(* Logix 5000 project; controller MV vendor 1 type 14 code 217 rev 31.11; software revision 31.00; part 41 of 53 *)
(* tags used below, declared in another part *)
   CurrentTime : DateTime;
   MV_B100 : INT[255];   // AT FLAGS
   MV_DayOfWeek : DINT;
   MV_F8 : REAL[20];
   MV_GasAvailable : BOOL;
   MV_MV10_CV1 : PlantItem;   // MV10_CV1
   MV_MV11_CV1 : PlantItem;   // MV11_CV1
   MV_MV12_CV1 : PlantItem;   // MV12_CV1
   MV_MV13_CV1 : PlantItem;   // MV13_CV1
   MV_MV14_CV1 : PlantItem;   // MV14_CV1
   MV_MV15_CV1 : PlantItem;   // MV15_CV1
   MV_MV16_CV1 : PlantItem;   // MV16_CV1
   MV_MV17_CV1 : PlantItem;   // MV17_CV1
   MV_MV18_CV1 : PlantItem;   // MV18_CV1
   MV_MV19_CV1 : PlantItem;   // MV19_CV1
   MV_MV1_CV1 : PlantItem;   // MV1_CV1
   MV_MV20_CV1 : PlantItem;   // MV20_CV1
   MV_MV21_CV1 : PlantItem;   // MV21_CV1
   MV_MV22_CV1 : PlantItem;   // MV22_CV1
   MV_MV23_CV1 : PlantItem;   // MV23_CV1
   MV_MV2_CV1 : PlantItem;   // MV2_CV1
   MV_MV30_CV1 : PlantItem;   // MV30_CV1
   MV_MV31_CV1 : PlantItem;   // MV31_CV1
   MV_MV32_CV1 : PlantItem;   // MV32_CV1
   MV_MV33_CV1 : PlantItem;   // MV33_CV1
   MV_MV34_CV1 : PlantItem;   // MV34_CV1
   MV_MV35_CV1 : PlantItem;   // MV35_CV1
   MV_MV36_AV01 : PlantItem;   // MV36_AV01
   MV_MV37_AV01 : PlantItem;   // MV37_AV01
   MV_MV38_AV01 : PlantItem;   // MV38_AV01
   MV_MV39_AV01 : PlantItem;   // MV39_AV01
   MV_MV3_CV1 : PlantItem;   // MV3_CV1
   MV_MV40_AV01 : PlantItem;   // MV40_AV01
   MV_MV41_AV01 : PlantItem;   // MV41_AV01
   MV_MV42_AV01 : PlantItem;   // MV42_AV01
   MV_MV43_AV01 : PlantItem;   // MV43_AV01
   MV_MV44_AV01 : PlantItem;   // MV44_AV01
   MV_MV45_AV01 : PlantItem;   // MV45_AV01
   MV_MV46_AV01 : PlantItem;   // MV46_AV01
   MV_MV47_AV01 : PlantItem;   // MV47_AV01
   MV_MV4_CV1 : PlantItem;   // MV4_CV1
   MV_MV5_CV1 : PlantItem;   // MV5_CV1
   MV_MV6_CV1 : PlantItem;   // MV6_CV1
   MV_MV7_CV1 : PlantItem;   // MV7_CV1
   MV_MV8_CV1 : PlantItem;   // MV8_CV1
   MV_MV9_CV1 : PlantItem;   // MV9_CV1
   MV_N101 : INT[255];   // AT INT Fermentation control integer workspace
   MV_N110 : INT[255];   // MV DATA 0 CURRENT FV DATA
   MV_N111 : INT[50];   // MV 1, CURRENT FV DATA
   MV_N112 : INT[50];   // MV 2, CURRENT FV DATA
   MV_N113 : INT[50];   // MV 3, CURRENT FV DATA
   MV_N114 : INT[50];   // MV 4, CURRENT FV DATA
   MV_N115 : INT[50];   // MV 5, CURRENT FV DATA
   MV_N116 : INT[50];   // MV 6, CURRENT FV DATA
   MV_N117 : INT[50];   // MV 7, CURRENT FV DATA
   MV_N118 : INT[50];   // MV 8, CURRENT FV DATA
   MV_N119 : INT[50];   // MV 9, CURRENT FV DATA
   MV_N12 : INT[255];   // SYS_PARMS System Parameter Fil e
   MV_N120 : INT[50];   // MV 10, CURRENT FV DATA
   MV_N121 : INT[50];   // MV 11, CURRENT FV DATA
   MV_N122 : INT[50];   // MV 12, CURRENT FV DATA
   MV_N123 : INT[50];   // MV 13, CURRENT FV DATA
   MV_N124 : INT[50];   // MV 14, CURRENT FV DATA
   MV_N125 : INT[50];   // MV 15, CURRENT FV DATA
   MV_N126 : INT[50];   // MV 16, CURRENT FV DATA
   MV_N127 : INT[50];   // MV 17, CURRENT FV DATA
   MV_N128 : INT[50];   // MV 18, CURRENT FV DATA
   MV_N129 : INT[50];   // MV 19, CURRENT FV DATA
   MV_N130 : INT[50];   // MV 30, CURRENT FV DATA
   MV_N131 : INT[50];   // MV 31, CURRENT FV DATA
   MV_N132 : INT[50];   // MV 32, CURRENT FV DATA
   MV_N133 : INT[50];   // MV 33, CURRENT FV DATA
   MV_N134 : INT[50];   // MV 34, CURRENT FV DATA
   MV_N135 : INT[50];   // MV 35, CURRENT FV DATA
   MV_N136 : INT[50];   // MV 20, CURRENT FV DATA
   MV_N137 : INT[50];   // MV 21, CURRENT FV DATA
   MV_N138 : INT[50];   // MV 22, CURRENT FV DATA
   MV_N139 : INT[50];   // MV 23, CURRENT FV DATA
   MV_N140 : INT[50];   // MV 36, CURRENT FV DATA
   MV_N141 : INT[50];   // MV 37, CURRENT FV DATA
   MV_N142 : INT[50];   // MV 38, CURRENT FV DATA
   MV_N143 : INT[50];   // MV 39, CURRENT FV DATA
   MV_N144 : INT[50];   // MV 40, CURRENT FV DATA
   MV_N145 : INT[50];   // MV 41, CURRENT FV DATA
   MV_N146 : INT[50];   // MV 42, CURRENT FV DATA
   MV_N147 : INT[50];   // MV 43, CURRENT FV DATA
   MV_N148 : INT[50];   // MV 44, CURRENT FV DATA
   MV_N149 : INT[50];   // MV 45, CURRENT FV DATA
   MV_N150 : INT[50];   // MV 36, CURRENT FV DATA
   MV_N151 : INT[50];   // MV 47, CURRENT FV DATA
   MV_SFile : INT[255];   // SLC Equivalent System File, So Original Code Can Remain
   temp : INT;
(* MV_Common, continued *)

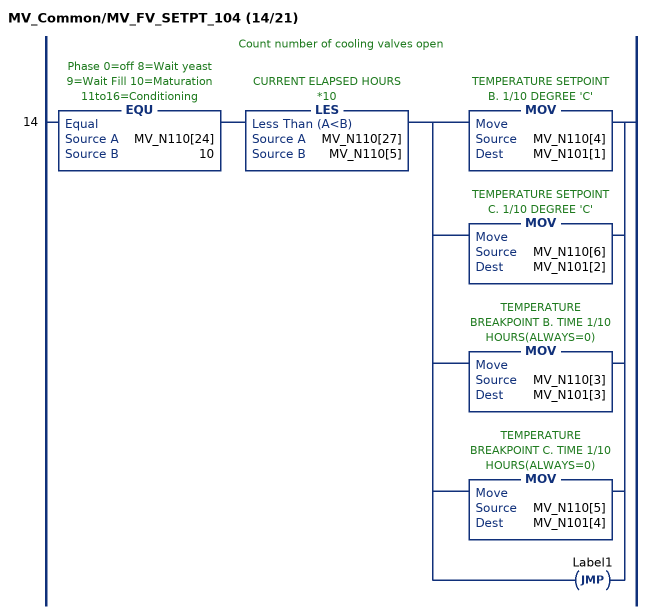
   [picture p954: MV_Common/MV_FV_SETPT_104 rungs 14-14]
   // Count number of cooling valves open
   14: EQU(MV_N110[24],10)LES(MV_N110[27],MV_N110[5])[MOV(MV_N110[4],MV_N101[1]) ,MOV(MV_N110[6],MV_N101[2]) ,MOV(MV_N110[3],MV_N101[3]) ,MOV(MV_N110[5],MV_N101[4]) ,JMP(Label1) ];
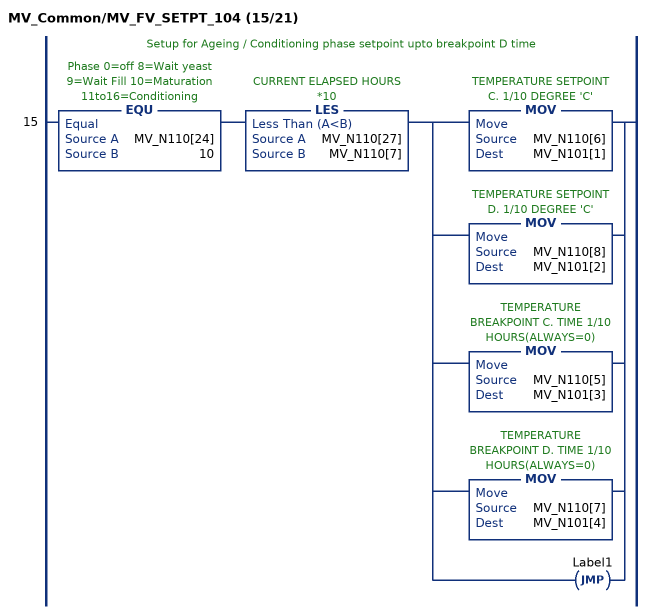
   // Setup for Ageing / Conditioning phase setpoint upto breakpoint D time
   15: EQU(MV_N110[24],10)LES(MV_N110[27],MV_N110[7])[MOV(MV_N110[6],MV_N101[1]) ,MOV(MV_N110[8],MV_N101[2]) ,MOV(MV_N110[5],MV_N101[3]) ,MOV(MV_N110[7],MV_N101[4]) ,JMP(Label1) ];
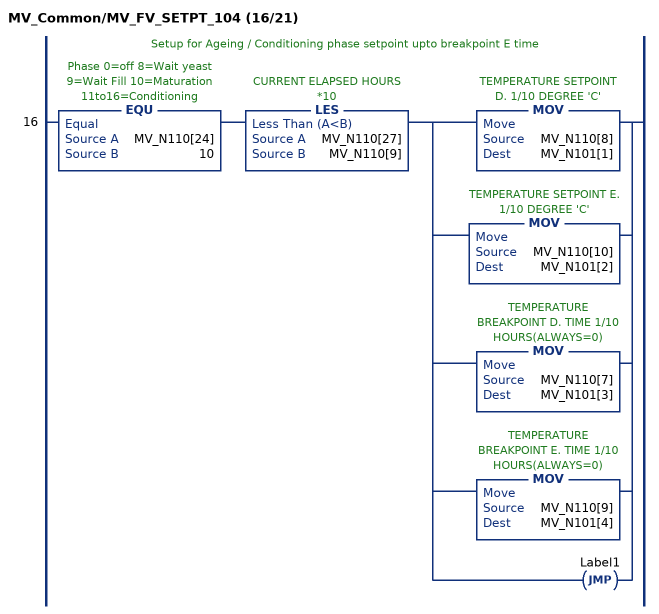
   // Setup for Ageing / Conditioning phase setpoint upto breakpoint E time
   16: EQU(MV_N110[24],10)LES(MV_N110[27],MV_N110[9])[MOV(MV_N110[8],MV_N101[1]) ,MOV(MV_N110[10],MV_N101[2]) ,MOV(MV_N110[7],MV_N101[3]) ,MOV(MV_N110[9],MV_N101[4]) ,JMP(Label1) ];
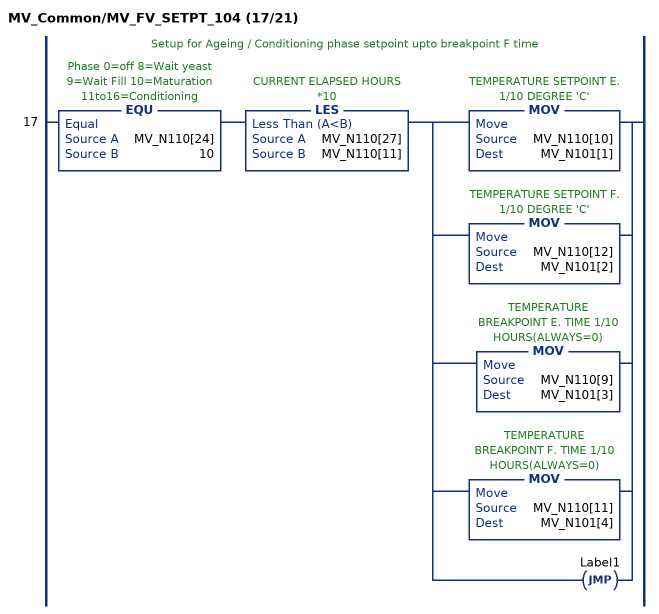
   // Setup for Ageing / Conditioning phase setpoint upto breakpoint F time
   17: EQU(MV_N110[24],10)LES(MV_N110[27],MV_N110[11])[MOV(MV_N110[10],MV_N101[1]) ,MOV(MV_N110[12],MV_N101[2]) ,MOV(MV_N110[9],MV_N101[3]) ,MOV(MV_N110[11],MV_N101[4]) ,JMP(Label1) ];
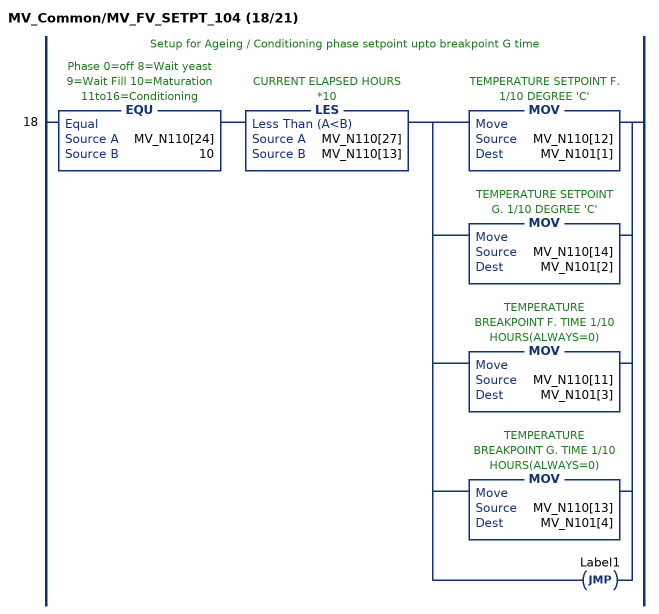
   // Setup for Ageing / Conditioning phase setpoint upto breakpoint G time
   18: EQU(MV_N110[24],10)LES(MV_N110[27],MV_N110[13])[MOV(MV_N110[12],MV_N101[1]) ,MOV(MV_N110[14],MV_N101[2]) ,MOV(MV_N110[11],MV_N101[3]) ,MOV(MV_N110[13],MV_N101[4]) ,JMP(Label1) ];
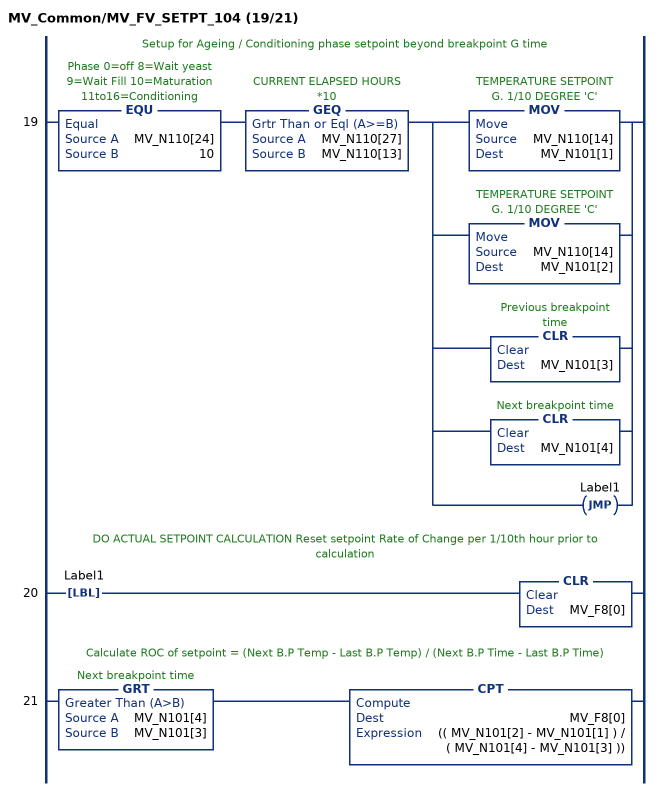
   // Setup for Ageing / Conditioning phase setpoint beyond breakpoint G time
   19: EQU(MV_N110[24],10)GEQ(MV_N110[27],MV_N110[13])[MOV(MV_N110[14],MV_N101[1]) ,MOV(MV_N110[14],MV_N101[2]) ,CLR(MV_N101[3]) ,CLR(MV_N101[4]) ,JMP(Label1) ];
   // DO ACTUAL SETPOINT CALCULATION Reset setpoint Rate of Change per 1/10th hour prior to calculation
   20: LBL(Label1)CLR(MV_F8[0]);
   // Calculate ROC of setpoint = (Next B.P Temp - Last B.P Temp) / (Next B.P Time - Last B.P Time)
   21: GRT(MV_N101[4],MV_N101[3])CPT(MV_F8[0],(( MV_N101[2] - MV_N101[1] ) / ( MV_N101[4] - MV_N101[3] )));
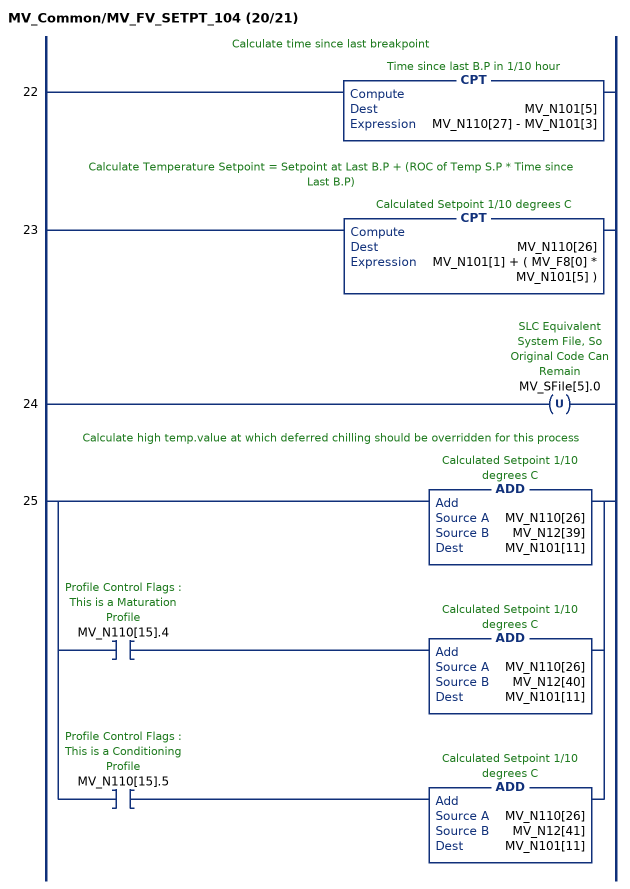
   // Calculate time since last breakpoint
   22: CPT(MV_N101[5],MV_N110[27] - MV_N101[3]);
   // Calculate Temperature Setpoint = Setpoint at Last B.P + (ROC of Temp S.P * Time since Last B.P)
   23: CPT(MV_N110[26],MV_N101[1] + ( MV_F8[0] * MV_N101[5] ));
   24: OTU(MV_SFile[5].0);
   // Calculate high temp.value at which deferred chilling should be overridden for this process
   25: [ADD(MV_N110[26],MV_N12[39],MV_N101[11]) ,XIC(MV_N110[15].4) ADD(MV_N110[26],MV_N12[40],MV_N101[11]) ,XIC(MV_N110[15].5) ADD(MV_N110[26],MV_N12[41],MV_N101[11]) ];
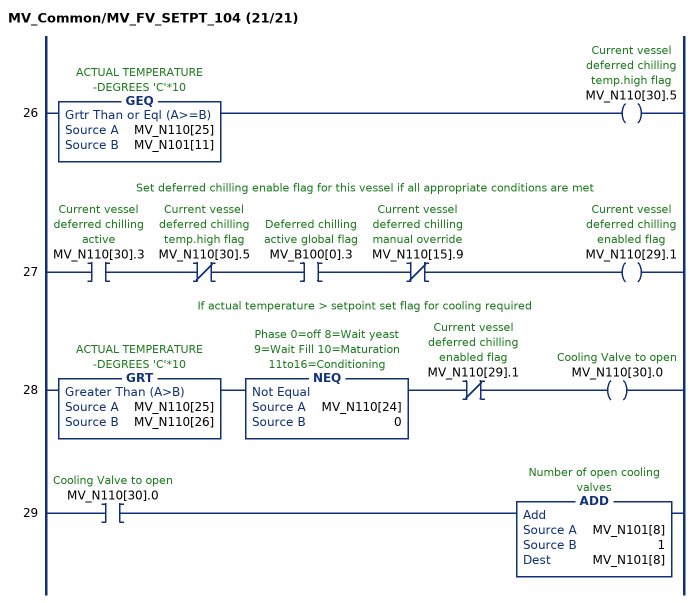
   26: GEQ(MV_N110[25],MV_N101[11])OTE(MV_N110[30].5);
   // Set deferred chilling enable flag for this vessel if all appropriate conditions are met
   27: XIC(MV_N110[30].3)XIO(MV_N110[30].5)XIC(MV_B100[0].3)XIO(MV_N110[15].9)OTE(MV_N110[29].1);
   // If actual temperature > setpoint set flag for cooling required
   28: GRT(MV_N110[25],MV_N110[26])NEQ(MV_N110[24],0)XIO(MV_N110[29].1)OTE(MV_N110[30].0);
   29: XIC(MV_N110[30].0)ADD(MV_N101[8],1,MV_N101[8]);
END_ROUTINE

ROUTINE MV_FV_VALVES_105   (* ladder *)
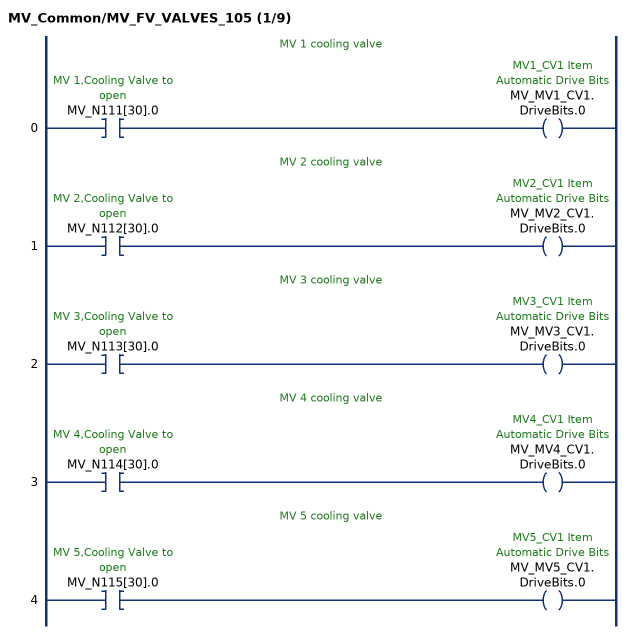
   // MV 1 cooling valve
   0: XIC(MV_N111[30].0)OTE(MV_MV1_CV1.DriveBits.0);
   // MV 2 cooling valve
   1: XIC(MV_N112[30].0)OTE(MV_MV2_CV1.DriveBits.0);
   // MV 3 cooling valve
   2: XIC(MV_N113[30].0)OTE(MV_MV3_CV1.DriveBits.0);
   // MV 4 cooling valve
   3: XIC(MV_N114[30].0)OTE(MV_MV4_CV1.DriveBits.0);
   // MV 5 cooling valve
   4: XIC(MV_N115[30].0)OTE(MV_MV5_CV1.DriveBits.0);
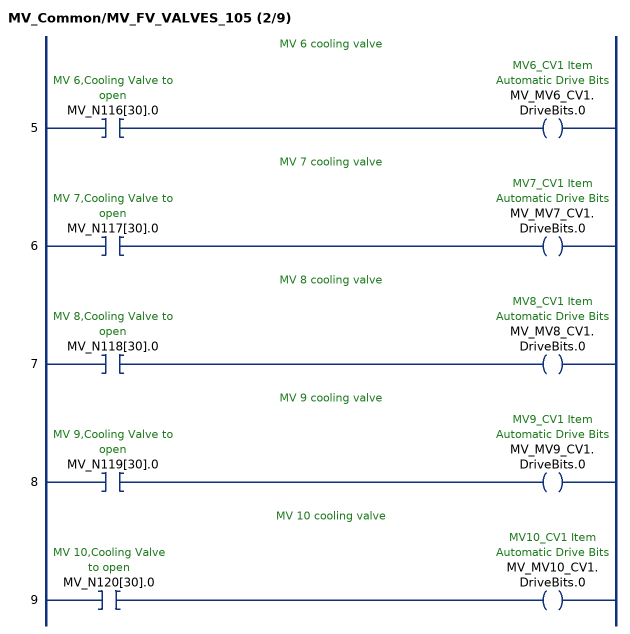
   // MV 6 cooling valve
   5: XIC(MV_N116[30].0)OTE(MV_MV6_CV1.DriveBits.0);
   // MV 7 cooling valve
   6: XIC(MV_N117[30].0)OTE(MV_MV7_CV1.DriveBits.0);
   // MV 8 cooling valve
   7: XIC(MV_N118[30].0)OTE(MV_MV8_CV1.DriveBits.0);
   // MV 9 cooling valve
   8: XIC(MV_N119[30].0)OTE(MV_MV9_CV1.DriveBits.0);
   // MV 10 cooling valve
   9: XIC(MV_N120[30].0)OTE(MV_MV10_CV1.DriveBits.0);
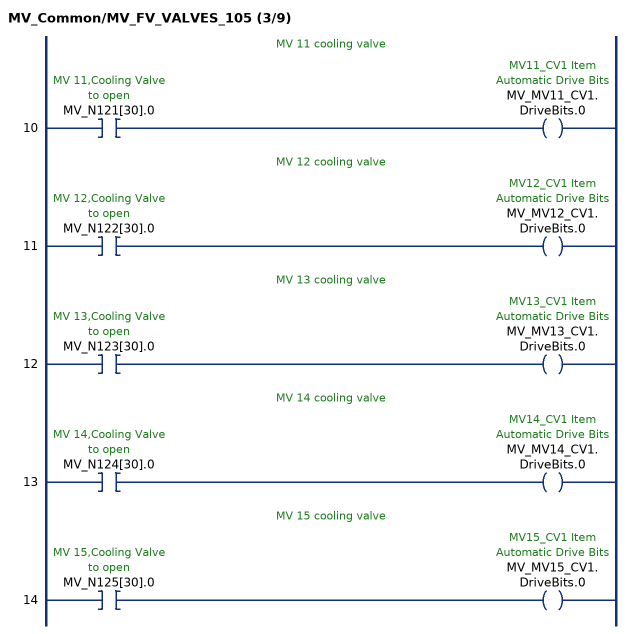
   // MV 11 cooling valve
   10: XIC(MV_N121[30].0)OTE(MV_MV11_CV1.DriveBits.0);
   // MV 12 cooling valve
   11: XIC(MV_N122[30].0)OTE(MV_MV12_CV1.DriveBits.0);
   // MV 13 cooling valve
   12: XIC(MV_N123[30].0)OTE(MV_MV13_CV1.DriveBits.0);
   // MV 14 cooling valve
   13: XIC(MV_N124[30].0)OTE(MV_MV14_CV1.DriveBits.0);
   // MV 15 cooling valve
   14: XIC(MV_N125[30].0)OTE(MV_MV15_CV1.DriveBits.0);
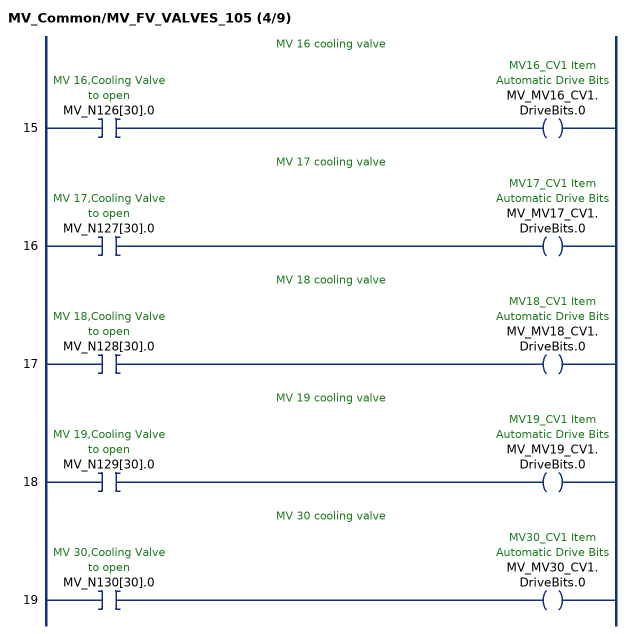
   // MV 16 cooling valve
   15: XIC(MV_N126[30].0)OTE(MV_MV16_CV1.DriveBits.0);
   // MV 17 cooling valve
   16: XIC(MV_N127[30].0)OTE(MV_MV17_CV1.DriveBits.0);
   // MV 18 cooling valve
   17: XIC(MV_N128[30].0)OTE(MV_MV18_CV1.DriveBits.0);
   // MV 19 cooling valve
   18: XIC(MV_N129[30].0)OTE(MV_MV19_CV1.DriveBits.0);
   // MV 30 cooling valve
   19: XIC(MV_N130[30].0)OTE(MV_MV30_CV1.DriveBits.0);
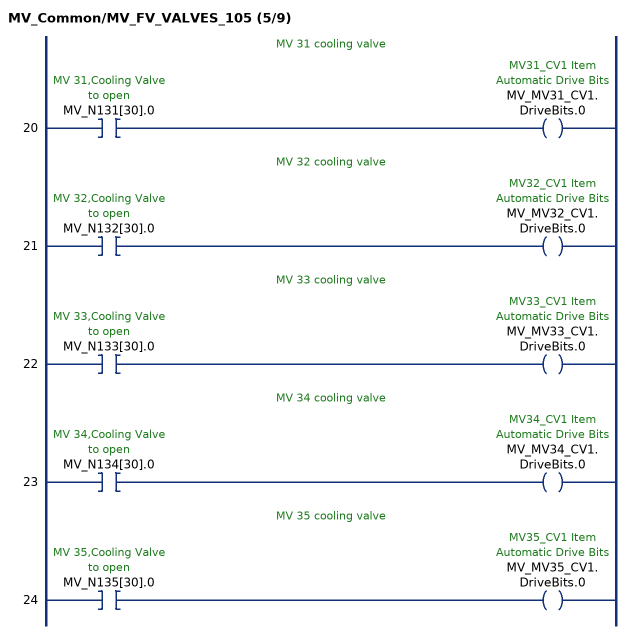
   // MV 31 cooling valve
   20: XIC(MV_N131[30].0)OTE(MV_MV31_CV1.DriveBits.0);
   // MV 32 cooling valve
   21: XIC(MV_N132[30].0)OTE(MV_MV32_CV1.DriveBits.0);
   // MV 33 cooling valve
   22: XIC(MV_N133[30].0)OTE(MV_MV33_CV1.DriveBits.0);
   // MV 34 cooling valve
   23: XIC(MV_N134[30].0)OTE(MV_MV34_CV1.DriveBits.0);
   // MV 35 cooling valve
   24: XIC(MV_N135[30].0)OTE(MV_MV35_CV1.DriveBits.0);
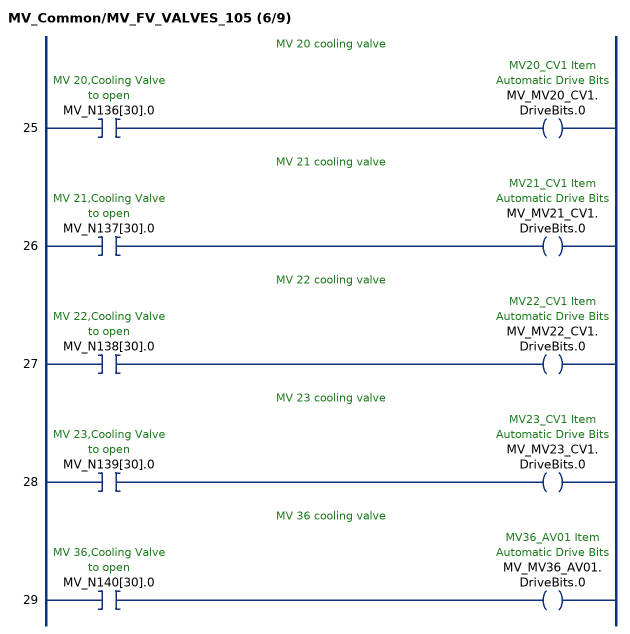
   // MV 20 cooling valve
   25: XIC(MV_N136[30].0)OTE(MV_MV20_CV1.DriveBits.0);
   // MV 21 cooling valve
   26: XIC(MV_N137[30].0)OTE(MV_MV21_CV1.DriveBits.0);
   // MV 22 cooling valve
   27: XIC(MV_N138[30].0)OTE(MV_MV22_CV1.DriveBits.0);
   // MV 23 cooling valve
   28: XIC(MV_N139[30].0)OTE(MV_MV23_CV1.DriveBits.0);
   // MV 36 cooling valve
   29: XIC(MV_N140[30].0)OTE(MV_MV36_AV01.DriveBits.0);
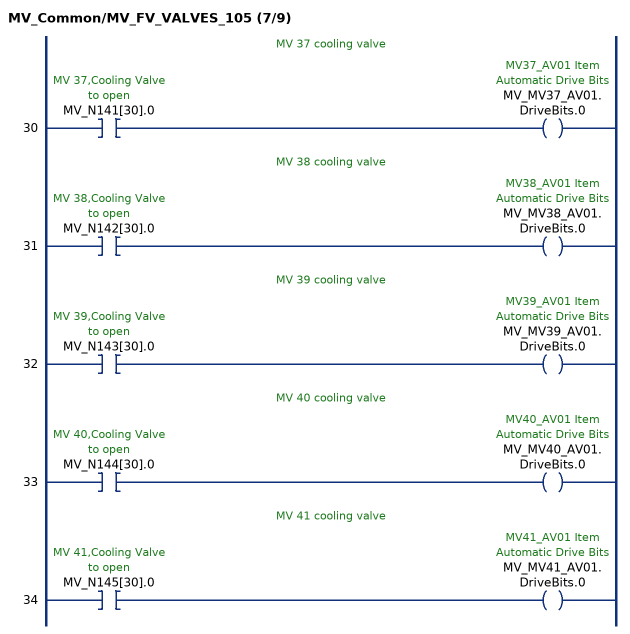
   // MV 37 cooling valve
   30: XIC(MV_N141[30].0)OTE(MV_MV37_AV01.DriveBits.0);
   // MV 38 cooling valve
   31: XIC(MV_N142[30].0)OTE(MV_MV38_AV01.DriveBits.0);
   // MV 39 cooling valve
   32: XIC(MV_N143[30].0)OTE(MV_MV39_AV01.DriveBits.0);
   // MV 40 cooling valve
   33: XIC(MV_N144[30].0)OTE(MV_MV40_AV01.DriveBits.0);
   // MV 41 cooling valve
   34: XIC(MV_N145[30].0)OTE(MV_MV41_AV01.DriveBits.0);
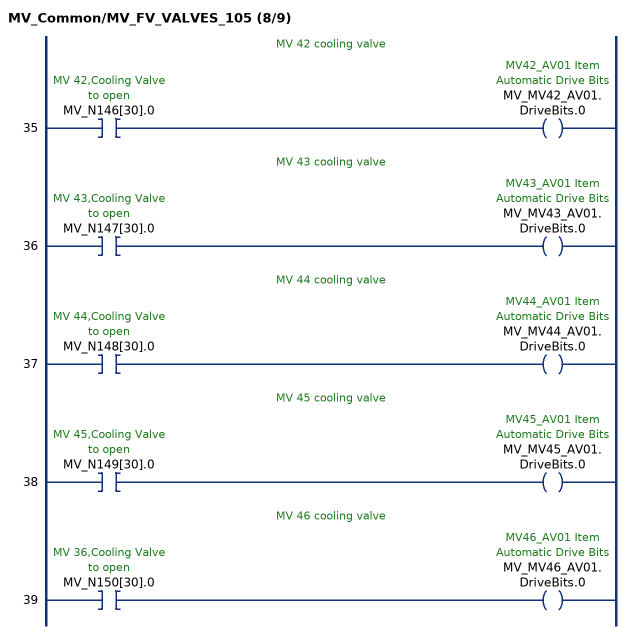
   // MV 42 cooling valve
   35: XIC(MV_N146[30].0)OTE(MV_MV42_AV01.DriveBits.0);
   // MV 43 cooling valve
   36: XIC(MV_N147[30].0)OTE(MV_MV43_AV01.DriveBits.0);
   // MV 44 cooling valve
   37: XIC(MV_N148[30].0)OTE(MV_MV44_AV01.DriveBits.0);
   // MV 45 cooling valve
   38: XIC(MV_N149[30].0)OTE(MV_MV45_AV01.DriveBits.0);
   // MV 46 cooling valve
   39: XIC(MV_N150[30].0)OTE(MV_MV46_AV01.DriveBits.0);
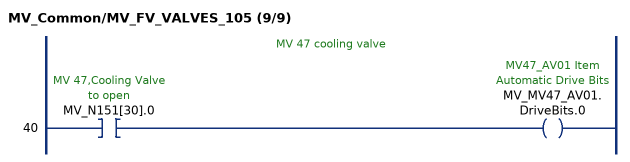
   // MV 47 cooling valve
   40: XIC(MV_N151[30].0)OTE(MV_MV47_AV01.DriveBits.0);
END_ROUTINE

ROUTINE MV_GAS_BLOCK   (* ladder *)
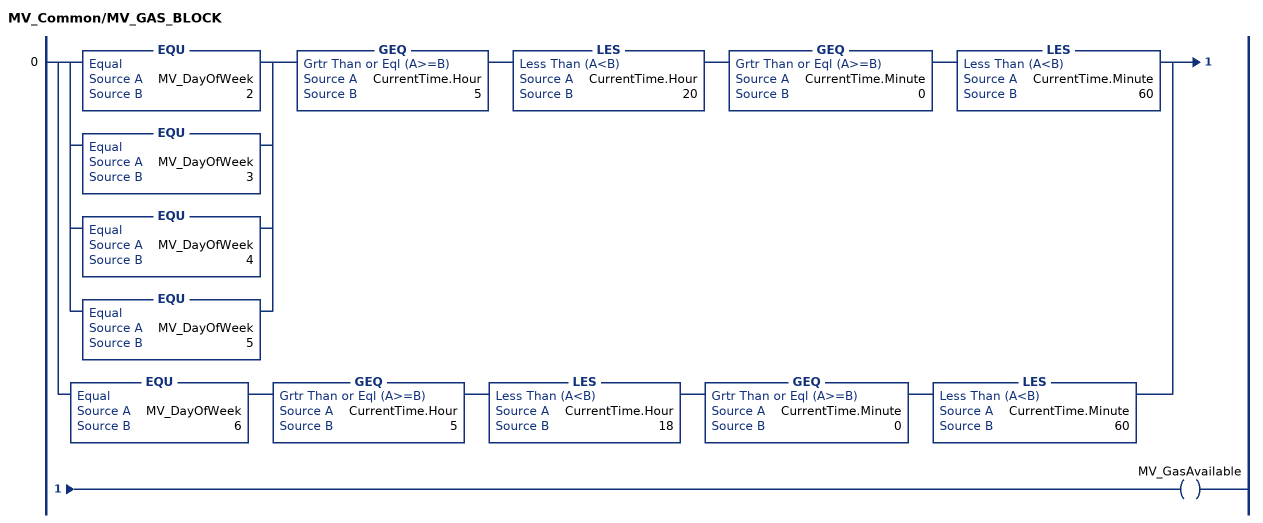
   0: [[EQU(MV_DayOfWeek,2) ,EQU(MV_DayOfWeek,3) ,EQU(MV_DayOfWeek,4) ,EQU(MV_DayOfWeek,5) ] GEQ(CurrentTime.Hour,5) LES(CurrentTime.Hour,20) GEQ(CurrentTime.Minute,0) LES(CurrentTime.Minute,60) ,EQU(MV_DayOfWeek,6) GEQ(CurrentTime.Hour,5) LES(CurrentTime.Hour,18) GEQ(CurrentTime.Minute,0) LES(CurrentTime.Minute,60) ]OTE(MV_GasAvailable);
END_ROUTINE
